(* Logix 5000 project; controller MV vendor 1 type 14 code 217 rev 31.11; software revision 31.00; part 19 of 53 *)
(* tags used below, declared in another part *)
   CheckTimeMask : INT;
   CWD : CHECKWORD_FLAGS;
   Delphi_Does_Eng_Func : BOOL;
   MC_CH1_DR1 : PlantItem;   // CH1_DR1
   MC_CH1_DR2 : PlantItem;   // CH1_DR2
   MC_CH1_DRAIN : PlantItem;   // CH1_DRAIN
   MC_CH1_R1R : PlantItem;   // CH1_R1R
   MC_CH1_R2R : PlantItem;   // CH1_R2R
   MC_CH1_R3R : PlantItem;   // CH1_R3R
   MC_CH1_R4 : PlantItem;   // CH1_R4
   MC_CH1_R4R : PlantItem;   // CH1_R4R
   MC_CH1_R5 : PlantItem;   // CH1_R5
   MC_CH1_R5R : PlantItem;   // CH1_R5R
   MC_CH1_R6 : PlantItem;   // CH1_R6
   MC_CH1_R6R : PlantItem;   // CH1_R6R
   MC_CH1_RR : PlantItem;   // CH1_RR
   MC_N255 : INT[255];   // CHECKWORDS Plant item checkword s
   TempChecktime : DINT;
(* MC_Common, continued *)

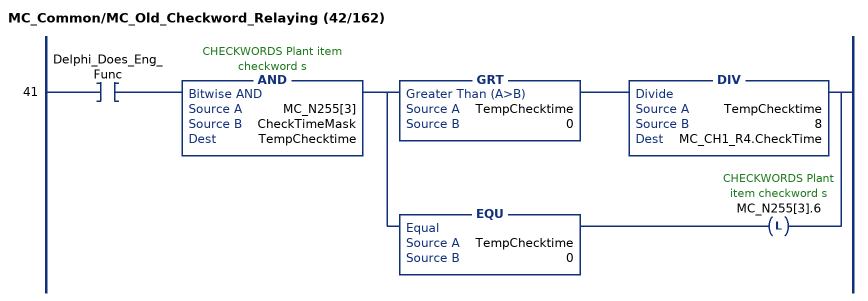
   [picture p312: MC_Common/MC_Old_Checkword_Relaying rungs 41-41]
   41: XIC(Delphi_Does_Eng_Func)AND(MC_N255[3],CheckTimeMask,TempChecktime)[GRT(TempChecktime,0) DIV(TempChecktime,8,MC_CH1_R4.CheckTime) ,EQU(TempChecktime,0) OTL(MC_N255[3].6) ];
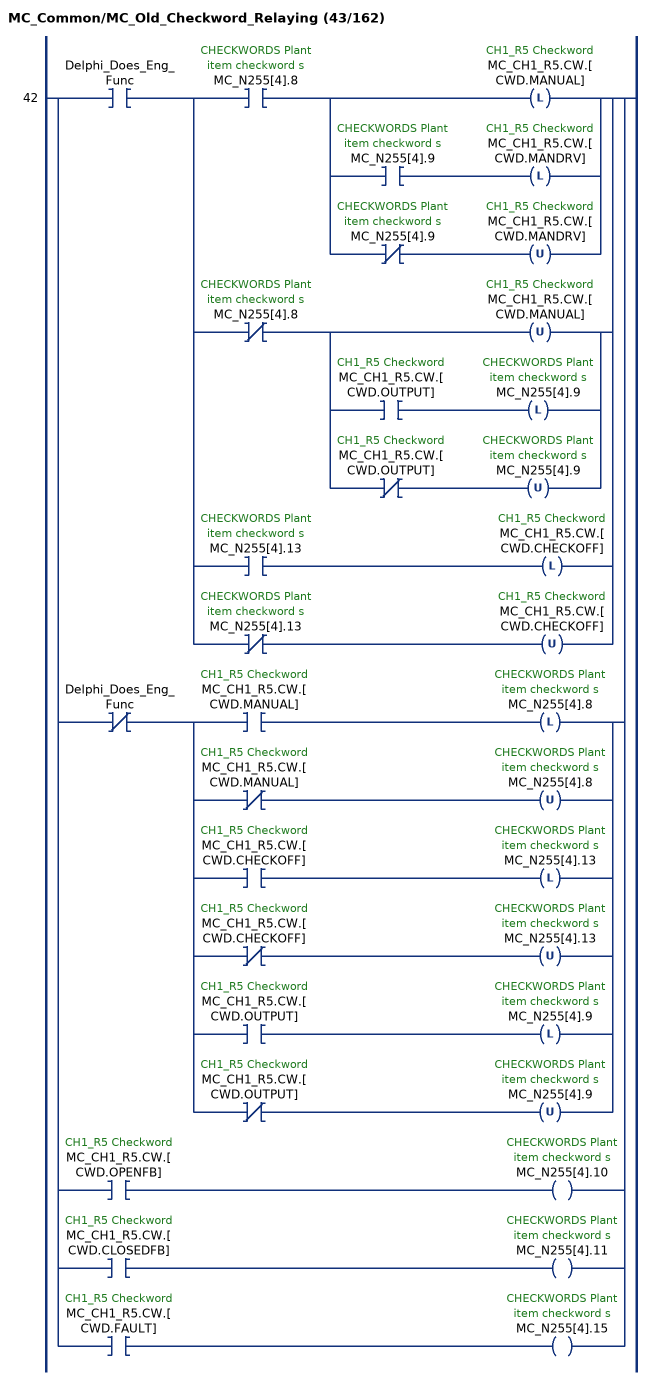
   42: [XIC(Delphi_Does_Eng_Func) [[XIC(MC_N255[4].8) [OTL(MC_CH1_R5.CW.[CWD.MANUAL]) ,XIC(MC_N255[4].9) OTL(MC_CH1_R5.CW.[CWD.MANDRV]) ,XIO(MC_N255[4].9) OTU(MC_CH1_R5.CW.[CWD.MANDRV]) ] ,XIO(MC_N255[4].8) [OTU(MC_CH1_R5.CW.[CWD.MANUAL]) ,[XIC(MC_CH1_R5.CW.[CWD.OUTPUT]) OTL(MC_N255[4].9) ,XIO(MC_CH1_R5.CW.[CWD.OUTPUT]) OTU(MC_N255[4].9) ] ] ] ,[XIC(MC_N255[4].13) OTL(MC_CH1_R5.CW.[CWD.CHECKOFF]) ,XIO(MC_N255[4].13) OTU(MC_CH1_R5.CW.[CWD.CHECKOFF]) ] ] ,XIO(Delphi_Does_Eng_Func) [[XIC(MC_CH1_R5.CW.[CWD.MANUAL]) OTL(MC_N255[4].8) ,XIO(MC_CH1_R5.CW.[CWD.MANUAL]) OTU(MC_N255[4].8) ] ,[XIC(MC_CH1_R5.CW.[CWD.CHECKOFF]) OTL(MC_N255[4].13) ,XIO(MC_CH1_R5.CW.[CWD.CHECKOFF]) OTU(MC_N255[4].13) ] ,[XIC(MC_CH1_R5.CW.[CWD.OUTPUT]) OTL(MC_N255[4].9) ,XIO(MC_CH1_R5.CW.[CWD.OUTPUT]) OTU(MC_N255[4].9) ] ] ,XIC(MC_CH1_R5.CW.[CWD.OPENFB]) OTE(MC_N255[4].10) ,XIC(MC_CH1_R5.CW.[CWD.CLOSEDFB]) OTE(MC_N255[4].11) ,XIC(MC_CH1_R5.CW.[CWD.FAULT]) OTE(MC_N255[4].15) ];
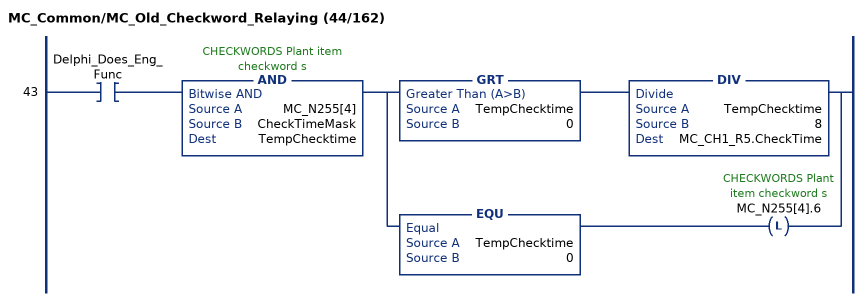
   43: XIC(Delphi_Does_Eng_Func)AND(MC_N255[4],CheckTimeMask,TempChecktime)[GRT(TempChecktime,0) DIV(TempChecktime,8,MC_CH1_R5.CheckTime) ,EQU(TempChecktime,0) OTL(MC_N255[4].6) ];
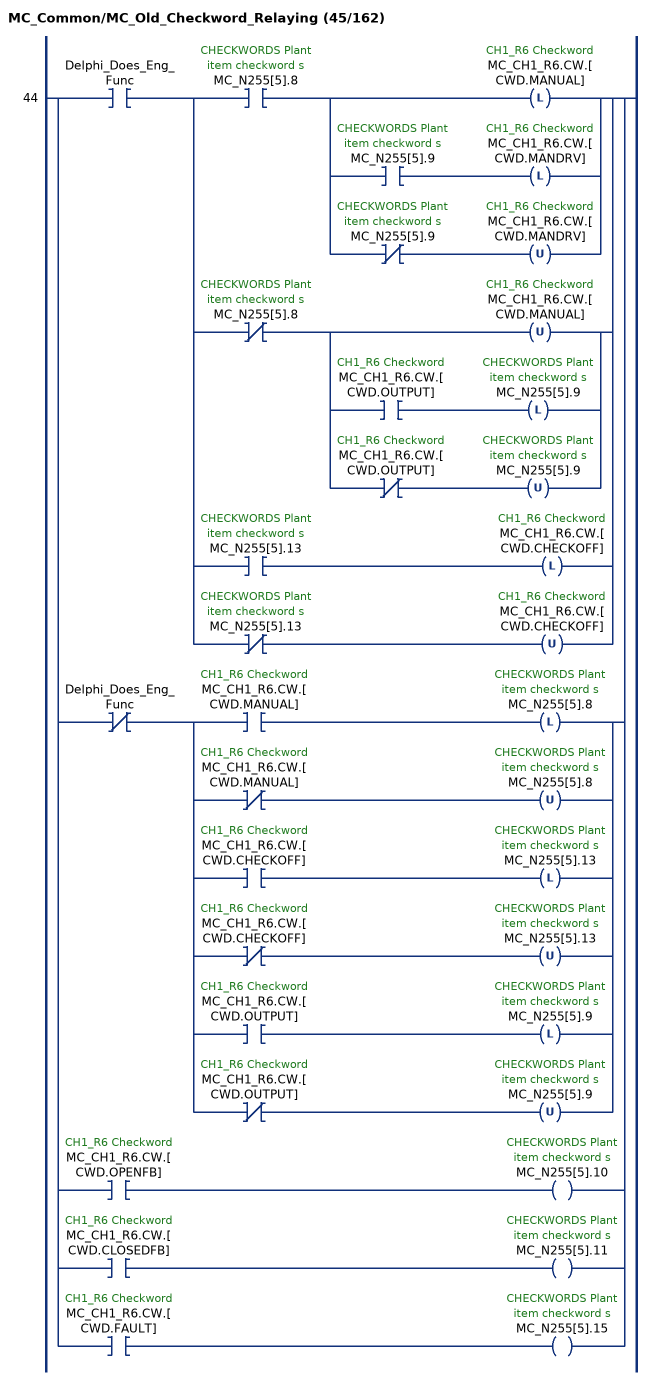
   44: [XIC(Delphi_Does_Eng_Func) [[XIC(MC_N255[5].8) [OTL(MC_CH1_R6.CW.[CWD.MANUAL]) ,XIC(MC_N255[5].9) OTL(MC_CH1_R6.CW.[CWD.MANDRV]) ,XIO(MC_N255[5].9) OTU(MC_CH1_R6.CW.[CWD.MANDRV]) ] ,XIO(MC_N255[5].8) [OTU(MC_CH1_R6.CW.[CWD.MANUAL]) ,[XIC(MC_CH1_R6.CW.[CWD.OUTPUT]) OTL(MC_N255[5].9) ,XIO(MC_CH1_R6.CW.[CWD.OUTPUT]) OTU(MC_N255[5].9) ] ] ] ,[XIC(MC_N255[5].13) OTL(MC_CH1_R6.CW.[CWD.CHECKOFF]) ,XIO(MC_N255[5].13) OTU(MC_CH1_R6.CW.[CWD.CHECKOFF]) ] ] ,XIO(Delphi_Does_Eng_Func) [[XIC(MC_CH1_R6.CW.[CWD.MANUAL]) OTL(MC_N255[5].8) ,XIO(MC_CH1_R6.CW.[CWD.MANUAL]) OTU(MC_N255[5].8) ] ,[XIC(MC_CH1_R6.CW.[CWD.CHECKOFF]) OTL(MC_N255[5].13) ,XIO(MC_CH1_R6.CW.[CWD.CHECKOFF]) OTU(MC_N255[5].13) ] ,[XIC(MC_CH1_R6.CW.[CWD.OUTPUT]) OTL(MC_N255[5].9) ,XIO(MC_CH1_R6.CW.[CWD.OUTPUT]) OTU(MC_N255[5].9) ] ] ,XIC(MC_CH1_R6.CW.[CWD.OPENFB]) OTE(MC_N255[5].10) ,XIC(MC_CH1_R6.CW.[CWD.CLOSEDFB]) OTE(MC_N255[5].11) ,XIC(MC_CH1_R6.CW.[CWD.FAULT]) OTE(MC_N255[5].15) ];
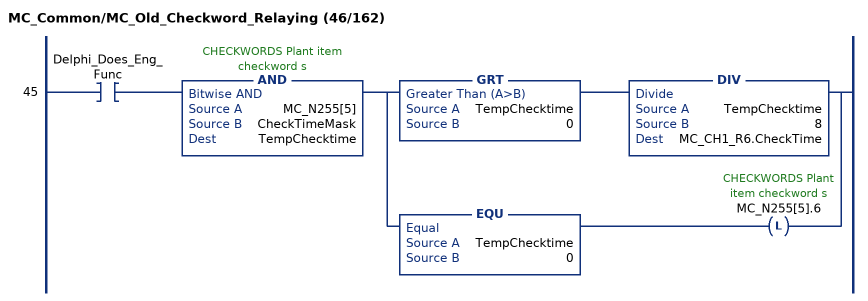
   45: XIC(Delphi_Does_Eng_Func)AND(MC_N255[5],CheckTimeMask,TempChecktime)[GRT(TempChecktime,0) DIV(TempChecktime,8,MC_CH1_R6.CheckTime) ,EQU(TempChecktime,0) OTL(MC_N255[5].6) ];
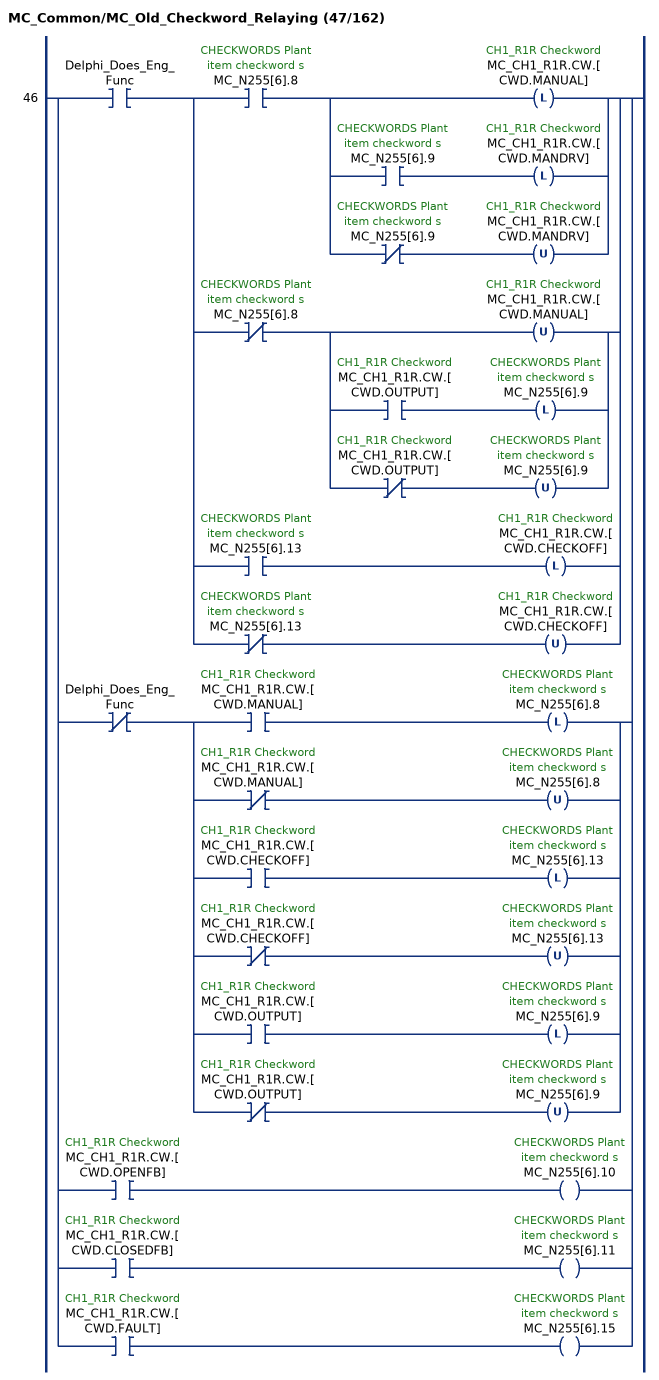
   46: [XIC(Delphi_Does_Eng_Func) [[XIC(MC_N255[6].8) [OTL(MC_CH1_R1R.CW.[CWD.MANUAL]) ,XIC(MC_N255[6].9) OTL(MC_CH1_R1R.CW.[CWD.MANDRV]) ,XIO(MC_N255[6].9) OTU(MC_CH1_R1R.CW.[CWD.MANDRV]) ] ,XIO(MC_N255[6].8) [OTU(MC_CH1_R1R.CW.[CWD.MANUAL]) ,[XIC(MC_CH1_R1R.CW.[CWD.OUTPUT]) OTL(MC_N255[6].9) ,XIO(MC_CH1_R1R.CW.[CWD.OUTPUT]) OTU(MC_N255[6].9) ] ] ] ,[XIC(MC_N255[6].13) OTL(MC_CH1_R1R.CW.[CWD.CHECKOFF]) ,XIO(MC_N255[6].13) OTU(MC_CH1_R1R.CW.[CWD.CHECKOFF]) ] ] ,XIO(Delphi_Does_Eng_Func) [[XIC(MC_CH1_R1R.CW.[CWD.MANUAL]) OTL(MC_N255[6].8) ,XIO(MC_CH1_R1R.CW.[CWD.MANUAL]) OTU(MC_N255[6].8) ] ,[XIC(MC_CH1_R1R.CW.[CWD.CHECKOFF]) OTL(MC_N255[6].13) ,XIO(MC_CH1_R1R.CW.[CWD.CHECKOFF]) OTU(MC_N255[6].13) ] ,[XIC(MC_CH1_R1R.CW.[CWD.OUTPUT]) OTL(MC_N255[6].9) ,XIO(MC_CH1_R1R.CW.[CWD.OUTPUT]) OTU(MC_N255[6].9) ] ] ,XIC(MC_CH1_R1R.CW.[CWD.OPENFB]) OTE(MC_N255[6].10) ,XIC(MC_CH1_R1R.CW.[CWD.CLOSEDFB]) OTE(MC_N255[6].11) ,XIC(MC_CH1_R1R.CW.[CWD.FAULT]) OTE(MC_N255[6].15) ];
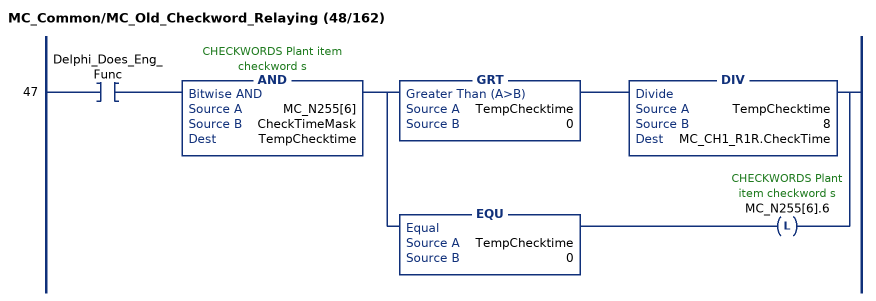
   47: XIC(Delphi_Does_Eng_Func)AND(MC_N255[6],CheckTimeMask,TempChecktime)[GRT(TempChecktime,0) DIV(TempChecktime,8,MC_CH1_R1R.CheckTime) ,EQU(TempChecktime,0) OTL(MC_N255[6].6) ];
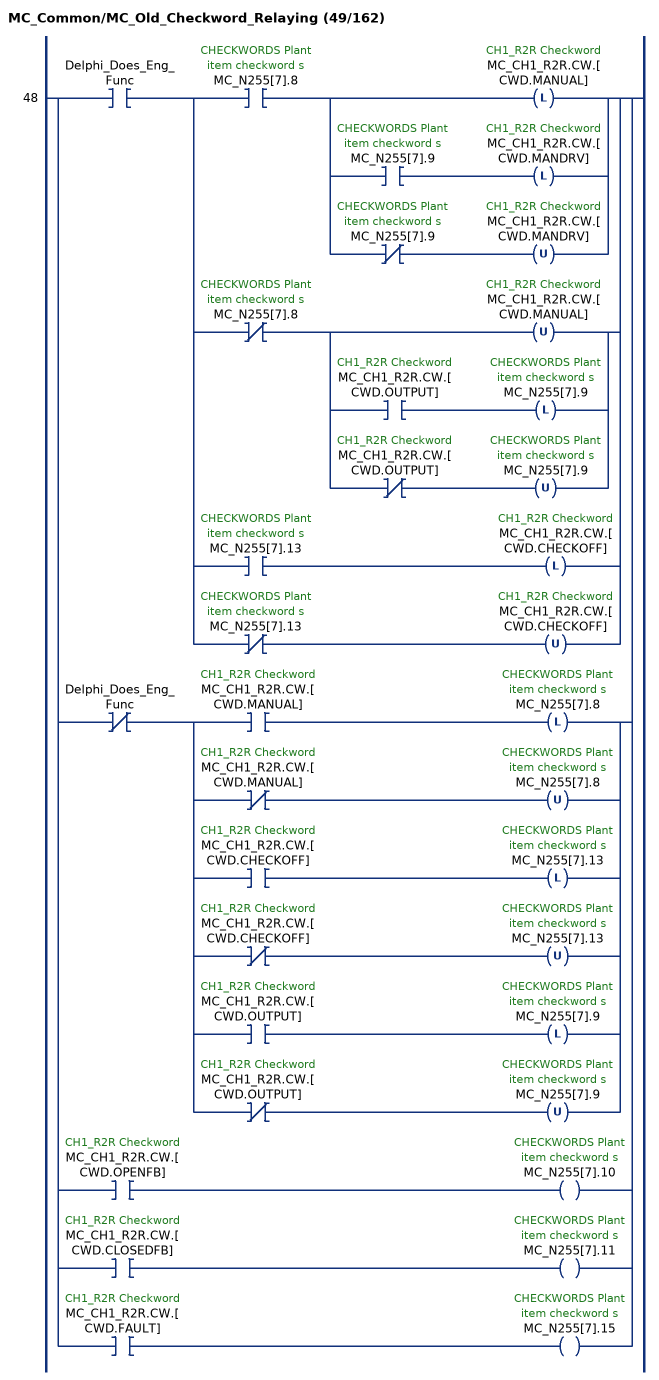
   48: [XIC(Delphi_Does_Eng_Func) [[XIC(MC_N255[7].8) [OTL(MC_CH1_R2R.CW.[CWD.MANUAL]) ,XIC(MC_N255[7].9) OTL(MC_CH1_R2R.CW.[CWD.MANDRV]) ,XIO(MC_N255[7].9) OTU(MC_CH1_R2R.CW.[CWD.MANDRV]) ] ,XIO(MC_N255[7].8) [OTU(MC_CH1_R2R.CW.[CWD.MANUAL]) ,[XIC(MC_CH1_R2R.CW.[CWD.OUTPUT]) OTL(MC_N255[7].9) ,XIO(MC_CH1_R2R.CW.[CWD.OUTPUT]) OTU(MC_N255[7].9) ] ] ] ,[XIC(MC_N255[7].13) OTL(MC_CH1_R2R.CW.[CWD.CHECKOFF]) ,XIO(MC_N255[7].13) OTU(MC_CH1_R2R.CW.[CWD.CHECKOFF]) ] ] ,XIO(Delphi_Does_Eng_Func) [[XIC(MC_CH1_R2R.CW.[CWD.MANUAL]) OTL(MC_N255[7].8) ,XIO(MC_CH1_R2R.CW.[CWD.MANUAL]) OTU(MC_N255[7].8) ] ,[XIC(MC_CH1_R2R.CW.[CWD.CHECKOFF]) OTL(MC_N255[7].13) ,XIO(MC_CH1_R2R.CW.[CWD.CHECKOFF]) OTU(MC_N255[7].13) ] ,[XIC(MC_CH1_R2R.CW.[CWD.OUTPUT]) OTL(MC_N255[7].9) ,XIO(MC_CH1_R2R.CW.[CWD.OUTPUT]) OTU(MC_N255[7].9) ] ] ,XIC(MC_CH1_R2R.CW.[CWD.OPENFB]) OTE(MC_N255[7].10) ,XIC(MC_CH1_R2R.CW.[CWD.CLOSEDFB]) OTE(MC_N255[7].11) ,XIC(MC_CH1_R2R.CW.[CWD.FAULT]) OTE(MC_N255[7].15) ];
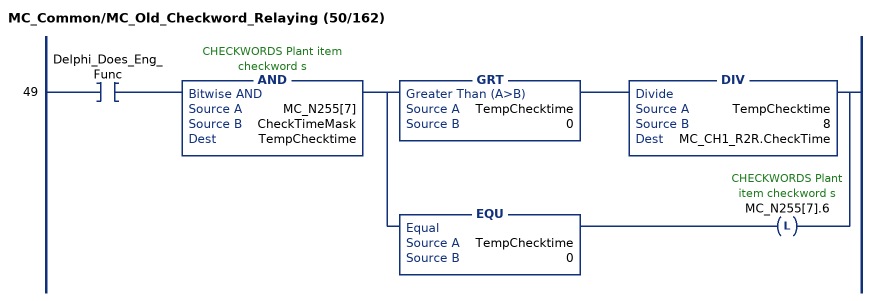
   49: XIC(Delphi_Does_Eng_Func)AND(MC_N255[7],CheckTimeMask,TempChecktime)[GRT(TempChecktime,0) DIV(TempChecktime,8,MC_CH1_R2R.CheckTime) ,EQU(TempChecktime,0) OTL(MC_N255[7].6) ];
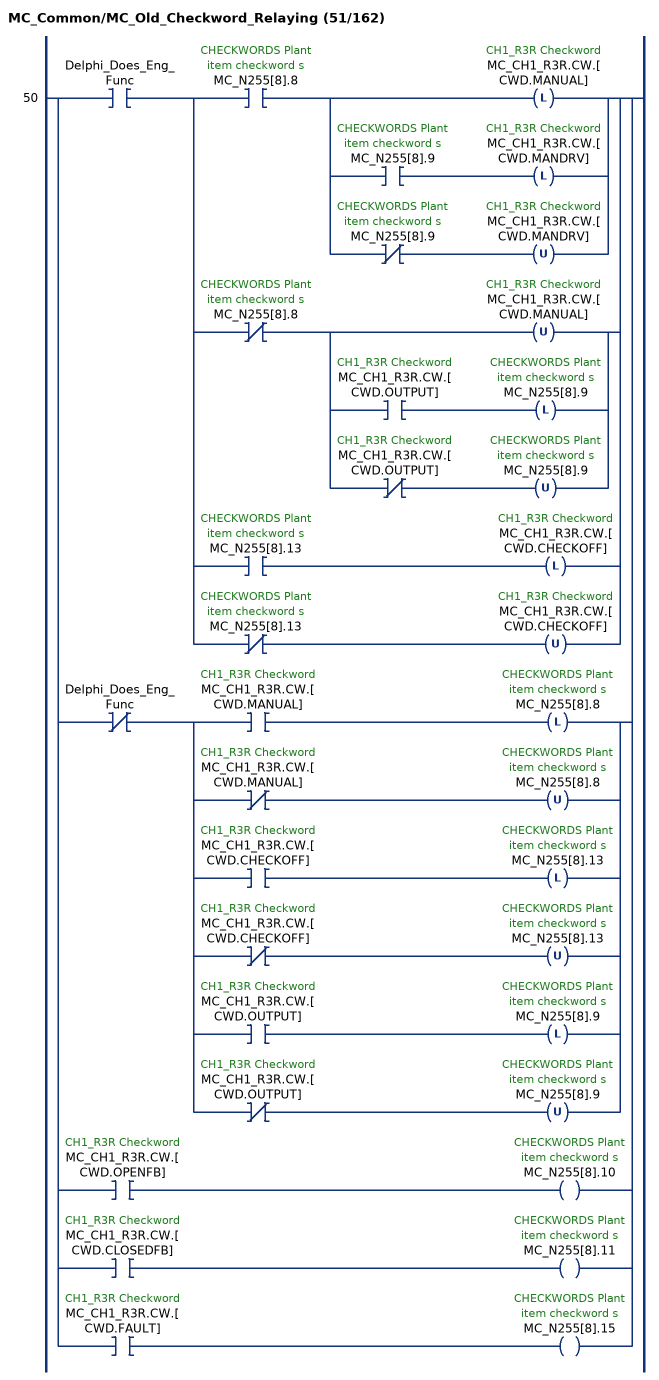
   50: [XIC(Delphi_Does_Eng_Func) [[XIC(MC_N255[8].8) [OTL(MC_CH1_R3R.CW.[CWD.MANUAL]) ,XIC(MC_N255[8].9) OTL(MC_CH1_R3R.CW.[CWD.MANDRV]) ,XIO(MC_N255[8].9) OTU(MC_CH1_R3R.CW.[CWD.MANDRV]) ] ,XIO(MC_N255[8].8) [OTU(MC_CH1_R3R.CW.[CWD.MANUAL]) ,[XIC(MC_CH1_R3R.CW.[CWD.OUTPUT]) OTL(MC_N255[8].9) ,XIO(MC_CH1_R3R.CW.[CWD.OUTPUT]) OTU(MC_N255[8].9) ] ] ] ,[XIC(MC_N255[8].13) OTL(MC_CH1_R3R.CW.[CWD.CHECKOFF]) ,XIO(MC_N255[8].13) OTU(MC_CH1_R3R.CW.[CWD.CHECKOFF]) ] ] ,XIO(Delphi_Does_Eng_Func) [[XIC(MC_CH1_R3R.CW.[CWD.MANUAL]) OTL(MC_N255[8].8) ,XIO(MC_CH1_R3R.CW.[CWD.MANUAL]) OTU(MC_N255[8].8) ] ,[XIC(MC_CH1_R3R.CW.[CWD.CHECKOFF]) OTL(MC_N255[8].13) ,XIO(MC_CH1_R3R.CW.[CWD.CHECKOFF]) OTU(MC_N255[8].13) ] ,[XIC(MC_CH1_R3R.CW.[CWD.OUTPUT]) OTL(MC_N255[8].9) ,XIO(MC_CH1_R3R.CW.[CWD.OUTPUT]) OTU(MC_N255[8].9) ] ] ,XIC(MC_CH1_R3R.CW.[CWD.OPENFB]) OTE(MC_N255[8].10) ,XIC(MC_CH1_R3R.CW.[CWD.CLOSEDFB]) OTE(MC_N255[8].11) ,XIC(MC_CH1_R3R.CW.[CWD.FAULT]) OTE(MC_N255[8].15) ];
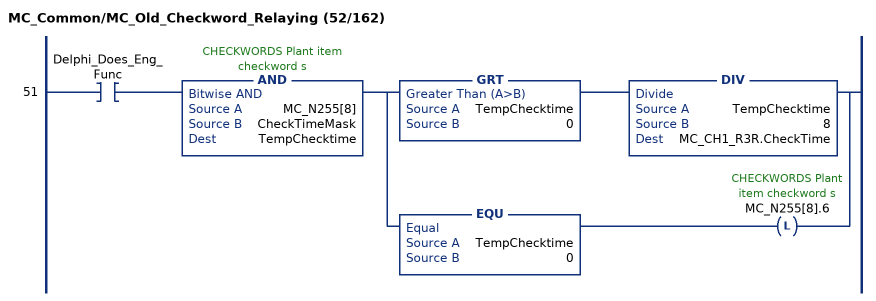
   51: XIC(Delphi_Does_Eng_Func)AND(MC_N255[8],CheckTimeMask,TempChecktime)[GRT(TempChecktime,0) DIV(TempChecktime,8,MC_CH1_R3R.CheckTime) ,EQU(TempChecktime,0) OTL(MC_N255[8].6) ];
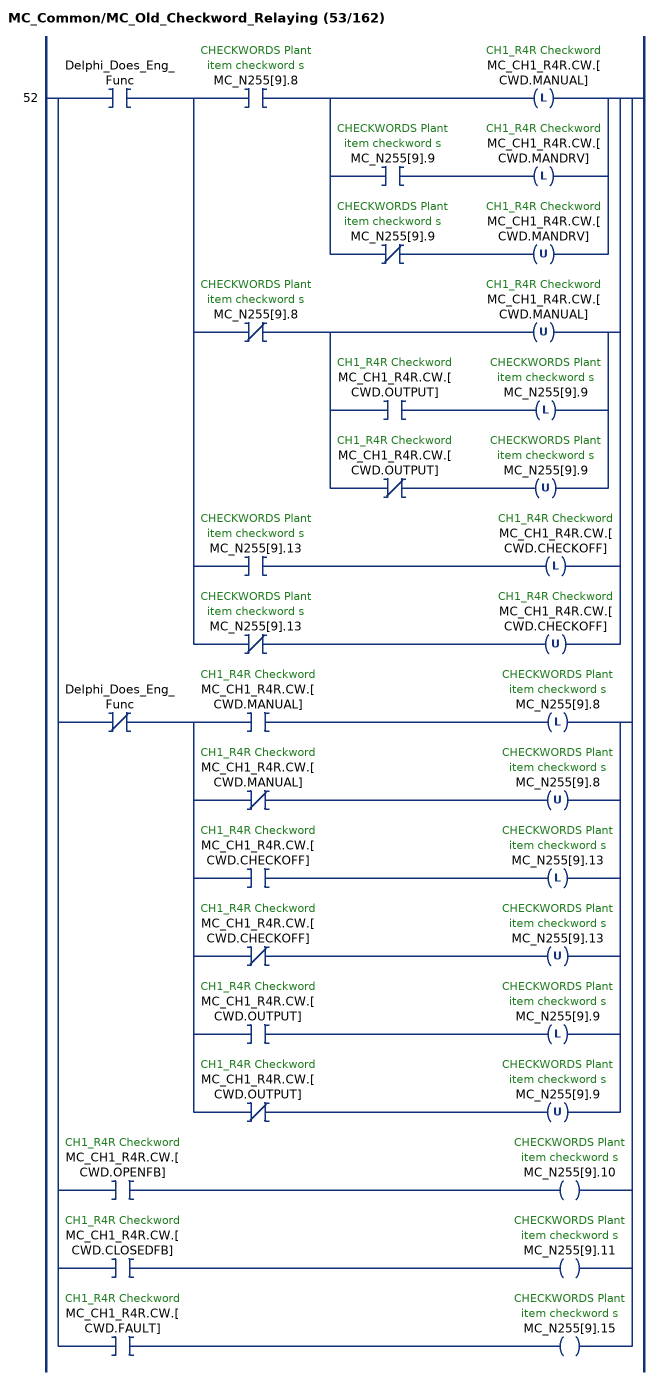
   52: [XIC(Delphi_Does_Eng_Func) [[XIC(MC_N255[9].8) [OTL(MC_CH1_R4R.CW.[CWD.MANUAL]) ,XIC(MC_N255[9].9) OTL(MC_CH1_R4R.CW.[CWD.MANDRV]) ,XIO(MC_N255[9].9) OTU(MC_CH1_R4R.CW.[CWD.MANDRV]) ] ,XIO(MC_N255[9].8) [OTU(MC_CH1_R4R.CW.[CWD.MANUAL]) ,[XIC(MC_CH1_R4R.CW.[CWD.OUTPUT]) OTL(MC_N255[9].9) ,XIO(MC_CH1_R4R.CW.[CWD.OUTPUT]) OTU(MC_N255[9].9) ] ] ] ,[XIC(MC_N255[9].13) OTL(MC_CH1_R4R.CW.[CWD.CHECKOFF]) ,XIO(MC_N255[9].13) OTU(MC_CH1_R4R.CW.[CWD.CHECKOFF]) ] ] ,XIO(Delphi_Does_Eng_Func) [[XIC(MC_CH1_R4R.CW.[CWD.MANUAL]) OTL(MC_N255[9].8) ,XIO(MC_CH1_R4R.CW.[CWD.MANUAL]) OTU(MC_N255[9].8) ] ,[XIC(MC_CH1_R4R.CW.[CWD.CHECKOFF]) OTL(MC_N255[9].13) ,XIO(MC_CH1_R4R.CW.[CWD.CHECKOFF]) OTU(MC_N255[9].13) ] ,[XIC(MC_CH1_R4R.CW.[CWD.OUTPUT]) OTL(MC_N255[9].9) ,XIO(MC_CH1_R4R.CW.[CWD.OUTPUT]) OTU(MC_N255[9].9) ] ] ,XIC(MC_CH1_R4R.CW.[CWD.OPENFB]) OTE(MC_N255[9].10) ,XIC(MC_CH1_R4R.CW.[CWD.CLOSEDFB]) OTE(MC_N255[9].11) ,XIC(MC_CH1_R4R.CW.[CWD.FAULT]) OTE(MC_N255[9].15) ];
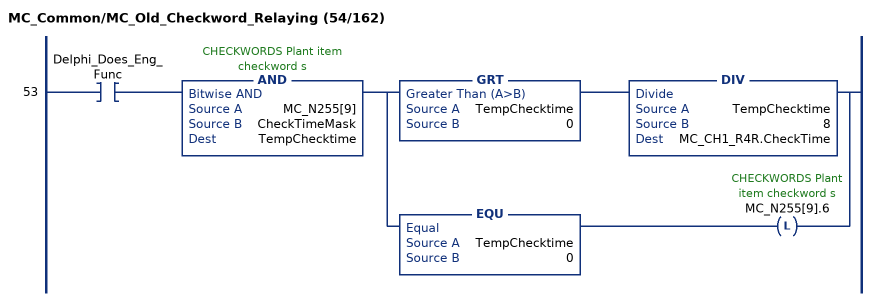
   53: XIC(Delphi_Does_Eng_Func)AND(MC_N255[9],CheckTimeMask,TempChecktime)[GRT(TempChecktime,0) DIV(TempChecktime,8,MC_CH1_R4R.CheckTime) ,EQU(TempChecktime,0) OTL(MC_N255[9].6) ];
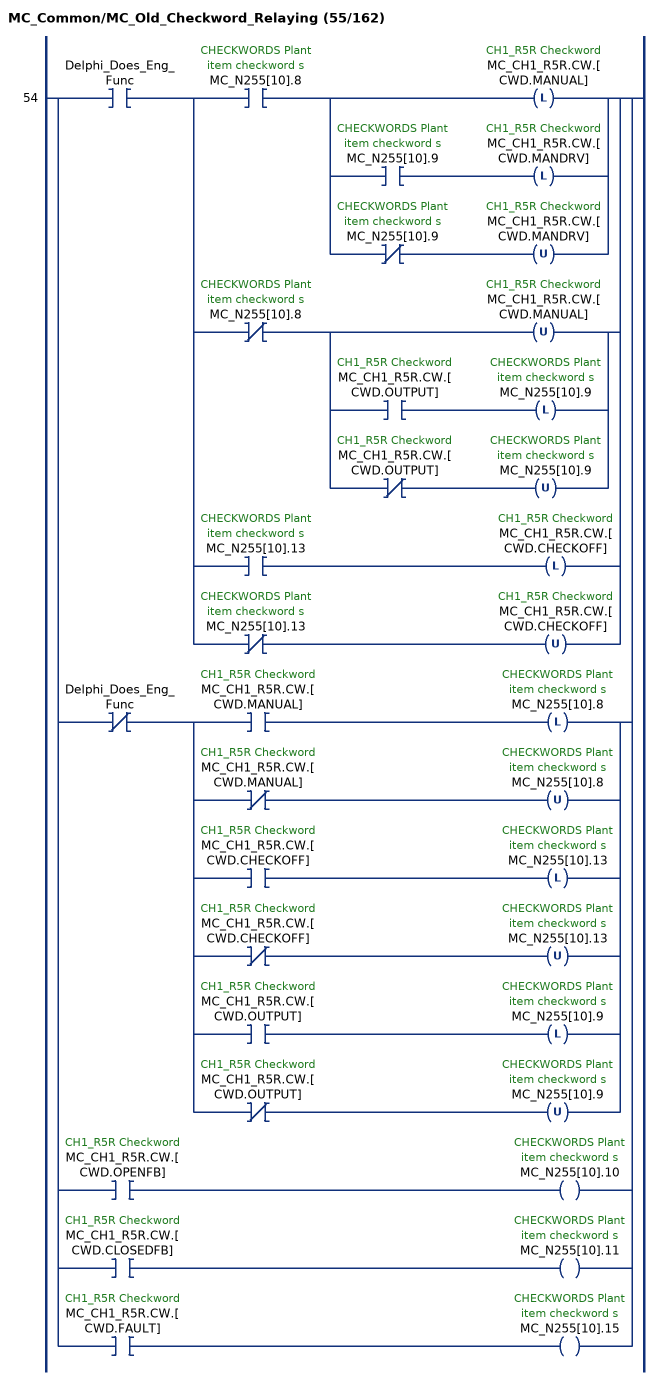
   54: [XIC(Delphi_Does_Eng_Func) [[XIC(MC_N255[10].8) [OTL(MC_CH1_R5R.CW.[CWD.MANUAL]) ,XIC(MC_N255[10].9) OTL(MC_CH1_R5R.CW.[CWD.MANDRV]) ,XIO(MC_N255[10].9) OTU(MC_CH1_R5R.CW.[CWD.MANDRV]) ] ,XIO(MC_N255[10].8) [OTU(MC_CH1_R5R.CW.[CWD.MANUAL]) ,[XIC(MC_CH1_R5R.CW.[CWD.OUTPUT]) OTL(MC_N255[10].9) ,XIO(MC_CH1_R5R.CW.[CWD.OUTPUT]) OTU(MC_N255[10].9) ] ] ] ,[XIC(MC_N255[10].13) OTL(MC_CH1_R5R.CW.[CWD.CHECKOFF]) ,XIO(MC_N255[10].13) OTU(MC_CH1_R5R.CW.[CWD.CHECKOFF]) ] ] ,XIO(Delphi_Does_Eng_Func) [[XIC(MC_CH1_R5R.CW.[CWD.MANUAL]) OTL(MC_N255[10].8) ,XIO(MC_CH1_R5R.CW.[CWD.MANUAL]) OTU(MC_N255[10].8) ] ,[XIC(MC_CH1_R5R.CW.[CWD.CHECKOFF]) OTL(MC_N255[10].13) ,XIO(MC_CH1_R5R.CW.[CWD.CHECKOFF]) OTU(MC_N255[10].13) ] ,[XIC(MC_CH1_R5R.CW.[CWD.OUTPUT]) OTL(MC_N255[10].9) ,XIO(MC_CH1_R5R.CW.[CWD.OUTPUT]) OTU(MC_N255[10].9) ] ] ,XIC(MC_CH1_R5R.CW.[CWD.OPENFB]) OTE(MC_N255[10].10) ,XIC(MC_CH1_R5R.CW.[CWD.CLOSEDFB]) OTE(MC_N255[10].11) ,XIC(MC_CH1_R5R.CW.[CWD.FAULT]) OTE(MC_N255[10].15) ];
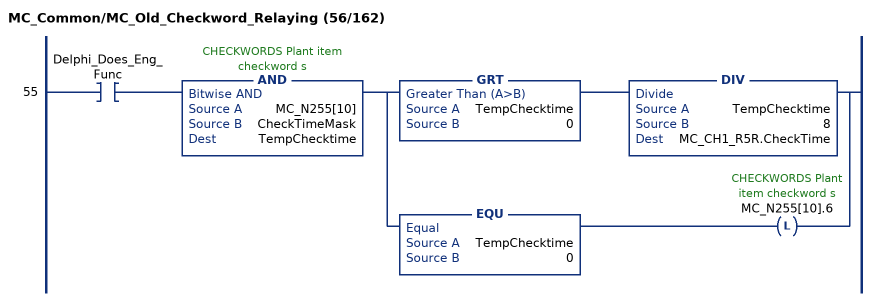
   55: XIC(Delphi_Does_Eng_Func)AND(MC_N255[10],CheckTimeMask,TempChecktime)[GRT(TempChecktime,0) DIV(TempChecktime,8,MC_CH1_R5R.CheckTime) ,EQU(TempChecktime,0) OTL(MC_N255[10].6) ];
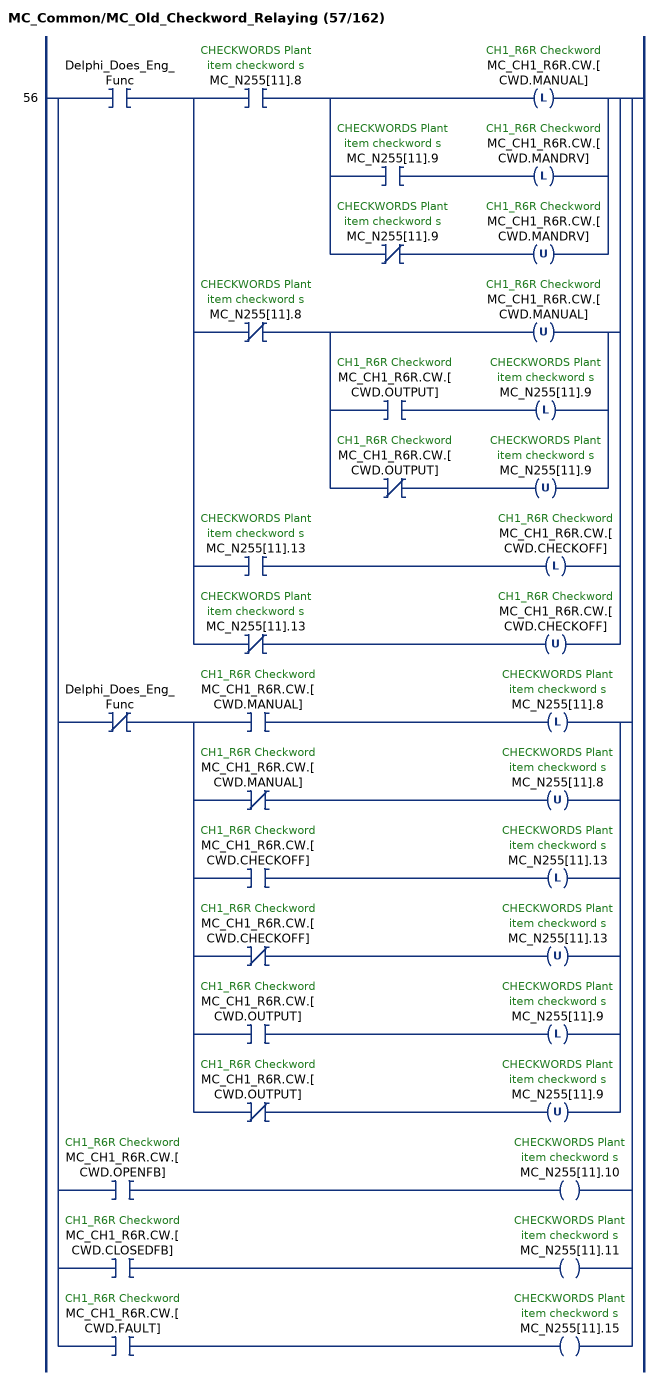
   56: [XIC(Delphi_Does_Eng_Func) [[XIC(MC_N255[11].8) [OTL(MC_CH1_R6R.CW.[CWD.MANUAL]) ,XIC(MC_N255[11].9) OTL(MC_CH1_R6R.CW.[CWD.MANDRV]) ,XIO(MC_N255[11].9) OTU(MC_CH1_R6R.CW.[CWD.MANDRV]) ] ,XIO(MC_N255[11].8) [OTU(MC_CH1_R6R.CW.[CWD.MANUAL]) ,[XIC(MC_CH1_R6R.CW.[CWD.OUTPUT]) OTL(MC_N255[11].9) ,XIO(MC_CH1_R6R.CW.[CWD.OUTPUT]) OTU(MC_N255[11].9) ] ] ] ,[XIC(MC_N255[11].13) OTL(MC_CH1_R6R.CW.[CWD.CHECKOFF]) ,XIO(MC_N255[11].13) OTU(MC_CH1_R6R.CW.[CWD.CHECKOFF]) ] ] ,XIO(Delphi_Does_Eng_Func) [[XIC(MC_CH1_R6R.CW.[CWD.MANUAL]) OTL(MC_N255[11].8) ,XIO(MC_CH1_R6R.CW.[CWD.MANUAL]) OTU(MC_N255[11].8) ] ,[XIC(MC_CH1_R6R.CW.[CWD.CHECKOFF]) OTL(MC_N255[11].13) ,XIO(MC_CH1_R6R.CW.[CWD.CHECKOFF]) OTU(MC_N255[11].13) ] ,[XIC(MC_CH1_R6R.CW.[CWD.OUTPUT]) OTL(MC_N255[11].9) ,XIO(MC_CH1_R6R.CW.[CWD.OUTPUT]) OTU(MC_N255[11].9) ] ] ,XIC(MC_CH1_R6R.CW.[CWD.OPENFB]) OTE(MC_N255[11].10) ,XIC(MC_CH1_R6R.CW.[CWD.CLOSEDFB]) OTE(MC_N255[11].11) ,XIC(MC_CH1_R6R.CW.[CWD.FAULT]) OTE(MC_N255[11].15) ];
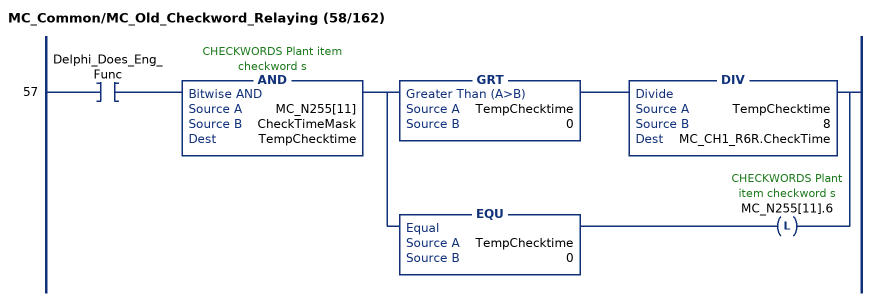
   57: XIC(Delphi_Does_Eng_Func)AND(MC_N255[11],CheckTimeMask,TempChecktime)[GRT(TempChecktime,0) DIV(TempChecktime,8,MC_CH1_R6R.CheckTime) ,EQU(TempChecktime,0) OTL(MC_N255[11].6) ];
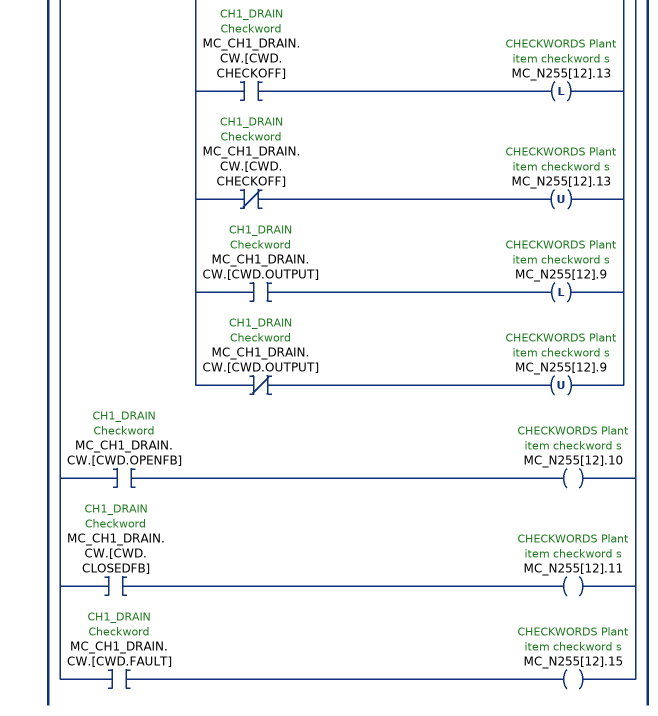
   58: [XIC(Delphi_Does_Eng_Func) [[XIC(MC_N255[12].8) [OTL(MC_CH1_DRAIN.CW.[CWD.MANUAL]) ,XIC(MC_N255[12].9) OTL(MC_CH1_DRAIN.CW.[CWD.MANDRV]) ,XIO(MC_N255[12].9) OTU(MC_CH1_DRAIN.CW.[CWD.MANDRV]) ] ,XIO(MC_N255[12].8) [OTU(MC_CH1_DRAIN.CW.[CWD.MANUAL]) ,[XIC(MC_CH1_DRAIN.CW.[CWD.OUTPUT]) OTL(MC_N255[12].9) ,XIO(MC_CH1_DRAIN.CW.[CWD.OUTPUT]) OTU(MC_N255[12].9) ] ] ] ,[XIC(MC_N255[12].13) OTL(MC_CH1_DRAIN.CW.[CWD.CHECKOFF]) ,XIO(MC_N255[12].13) OTU(MC_CH1_DRAIN.CW.[CWD.CHECKOFF]) ] ] ,XIO(Delphi_Does_Eng_Func) [[XIC(MC_CH1_DRAIN.CW.[CWD.MANUAL]) OTL(MC_N255[12].8) ,XIO(MC_CH1_DRAIN.CW.[CWD.MANUAL]) OTU(MC_N255[12].8) ] ,[XIC(MC_CH1_DRAIN.CW.[CWD.CHECKOFF]) OTL(MC_N255[12].13) ,XIO(MC_CH1_DRAIN.CW.[CWD.CHECKOFF]) OTU(MC_N255[12].13) ] ,[XIC(MC_CH1_DRAIN.CW.[CWD.OUTPUT]) OTL(MC_N255[12].9) ,XIO(MC_CH1_DRAIN.CW.[CWD.OUTPUT]) OTU(MC_N255[12].9) ] ] ,XIC(MC_CH1_DRAIN.CW.[CWD.OPENFB]) OTE(MC_N255[12].10) ,XIC(MC_CH1_DRAIN.CW.[CWD.CLOSEDFB]) OTE(MC_N255[12].11) ,XIC(MC_CH1_DRAIN.CW.[CWD.FAULT]) OTE(MC_N255[12].15) ];
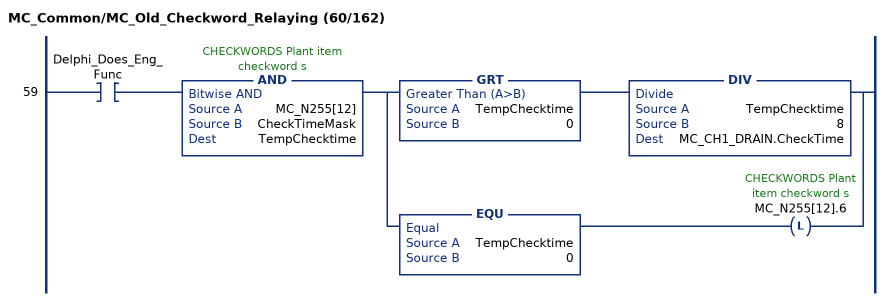
   59: XIC(Delphi_Does_Eng_Func)AND(MC_N255[12],CheckTimeMask,TempChecktime)[GRT(TempChecktime,0) DIV(TempChecktime,8,MC_CH1_DRAIN.CheckTime) ,EQU(TempChecktime,0) OTL(MC_N255[12].6) ];
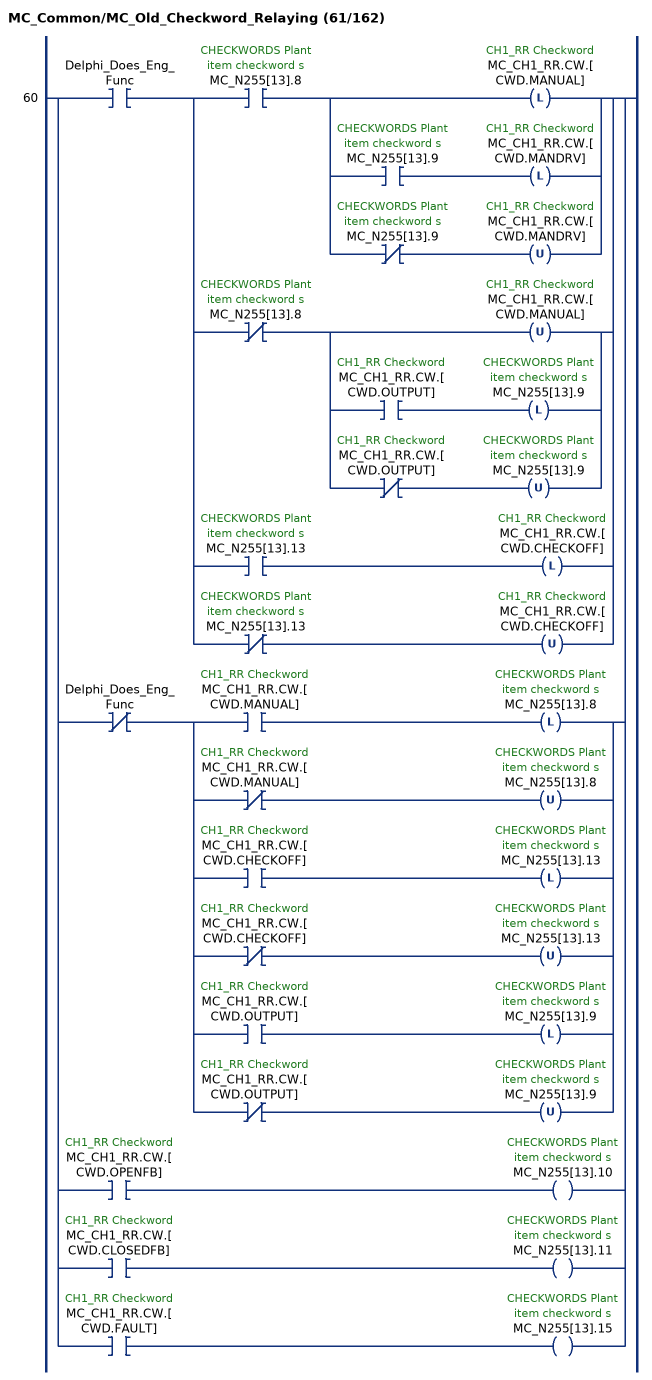
   60: [XIC(Delphi_Does_Eng_Func) [[XIC(MC_N255[13].8) [OTL(MC_CH1_RR.CW.[CWD.MANUAL]) ,XIC(MC_N255[13].9) OTL(MC_CH1_RR.CW.[CWD.MANDRV]) ,XIO(MC_N255[13].9) OTU(MC_CH1_RR.CW.[CWD.MANDRV]) ] ,XIO(MC_N255[13].8) [OTU(MC_CH1_RR.CW.[CWD.MANUAL]) ,[XIC(MC_CH1_RR.CW.[CWD.OUTPUT]) OTL(MC_N255[13].9) ,XIO(MC_CH1_RR.CW.[CWD.OUTPUT]) OTU(MC_N255[13].9) ] ] ] ,[XIC(MC_N255[13].13) OTL(MC_CH1_RR.CW.[CWD.CHECKOFF]) ,XIO(MC_N255[13].13) OTU(MC_CH1_RR.CW.[CWD.CHECKOFF]) ] ] ,XIO(Delphi_Does_Eng_Func) [[XIC(MC_CH1_RR.CW.[CWD.MANUAL]) OTL(MC_N255[13].8) ,XIO(MC_CH1_RR.CW.[CWD.MANUAL]) OTU(MC_N255[13].8) ] ,[XIC(MC_CH1_RR.CW.[CWD.CHECKOFF]) OTL(MC_N255[13].13) ,XIO(MC_CH1_RR.CW.[CWD.CHECKOFF]) OTU(MC_N255[13].13) ] ,[XIC(MC_CH1_RR.CW.[CWD.OUTPUT]) OTL(MC_N255[13].9) ,XIO(MC_CH1_RR.CW.[CWD.OUTPUT]) OTU(MC_N255[13].9) ] ] ,XIC(MC_CH1_RR.CW.[CWD.OPENFB]) OTE(MC_N255[13].10) ,XIC(MC_CH1_RR.CW.[CWD.CLOSEDFB]) OTE(MC_N255[13].11) ,XIC(MC_CH1_RR.CW.[CWD.FAULT]) OTE(MC_N255[13].15) ];
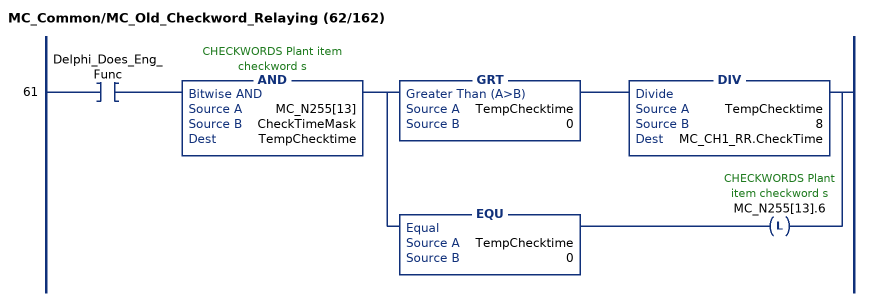
   61: XIC(Delphi_Does_Eng_Func)AND(MC_N255[13],CheckTimeMask,TempChecktime)[GRT(TempChecktime,0) DIV(TempChecktime,8,MC_CH1_RR.CheckTime) ,EQU(TempChecktime,0) OTL(MC_N255[13].6) ];
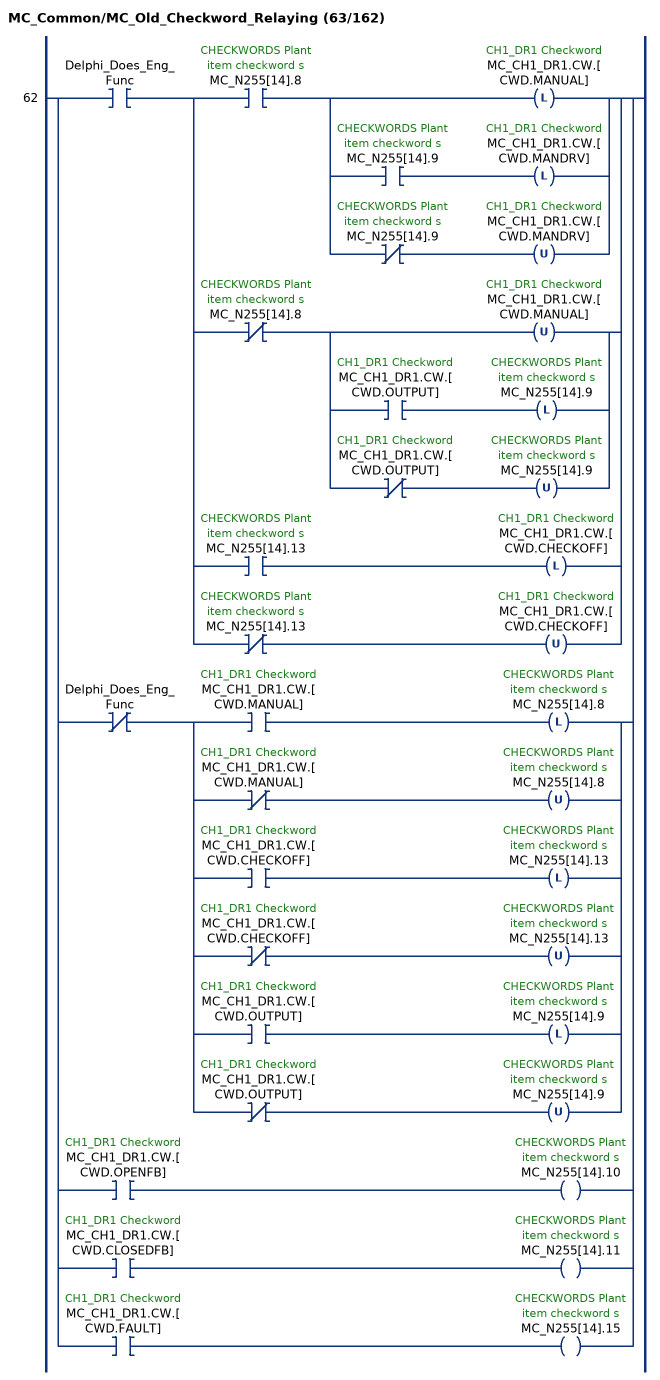
   62: [XIC(Delphi_Does_Eng_Func) [[XIC(MC_N255[14].8) [OTL(MC_CH1_DR1.CW.[CWD.MANUAL]) ,XIC(MC_N255[14].9) OTL(MC_CH1_DR1.CW.[CWD.MANDRV]) ,XIO(MC_N255[14].9) OTU(MC_CH1_DR1.CW.[CWD.MANDRV]) ] ,XIO(MC_N255[14].8) [OTU(MC_CH1_DR1.CW.[CWD.MANUAL]) ,[XIC(MC_CH1_DR1.CW.[CWD.OUTPUT]) OTL(MC_N255[14].9) ,XIO(MC_CH1_DR1.CW.[CWD.OUTPUT]) OTU(MC_N255[14].9) ] ] ] ,[XIC(MC_N255[14].13) OTL(MC_CH1_DR1.CW.[CWD.CHECKOFF]) ,XIO(MC_N255[14].13) OTU(MC_CH1_DR1.CW.[CWD.CHECKOFF]) ] ] ,XIO(Delphi_Does_Eng_Func) [[XIC(MC_CH1_DR1.CW.[CWD.MANUAL]) OTL(MC_N255[14].8) ,XIO(MC_CH1_DR1.CW.[CWD.MANUAL]) OTU(MC_N255[14].8) ] ,[XIC(MC_CH1_DR1.CW.[CWD.CHECKOFF]) OTL(MC_N255[14].13) ,XIO(MC_CH1_DR1.CW.[CWD.CHECKOFF]) OTU(MC_N255[14].13) ] ,[XIC(MC_CH1_DR1.CW.[CWD.OUTPUT]) OTL(MC_N255[14].9) ,XIO(MC_CH1_DR1.CW.[CWD.OUTPUT]) OTU(MC_N255[14].9) ] ] ,XIC(MC_CH1_DR1.CW.[CWD.OPENFB]) OTE(MC_N255[14].10) ,XIC(MC_CH1_DR1.CW.[CWD.CLOSEDFB]) OTE(MC_N255[14].11) ,XIC(MC_CH1_DR1.CW.[CWD.FAULT]) OTE(MC_N255[14].15) ];
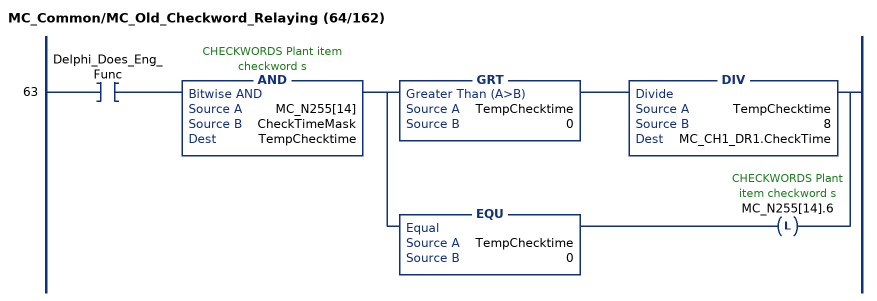
   63: XIC(Delphi_Does_Eng_Func)AND(MC_N255[14],CheckTimeMask,TempChecktime)[GRT(TempChecktime,0) DIV(TempChecktime,8,MC_CH1_DR1.CheckTime) ,EQU(TempChecktime,0) OTL(MC_N255[14].6) ];
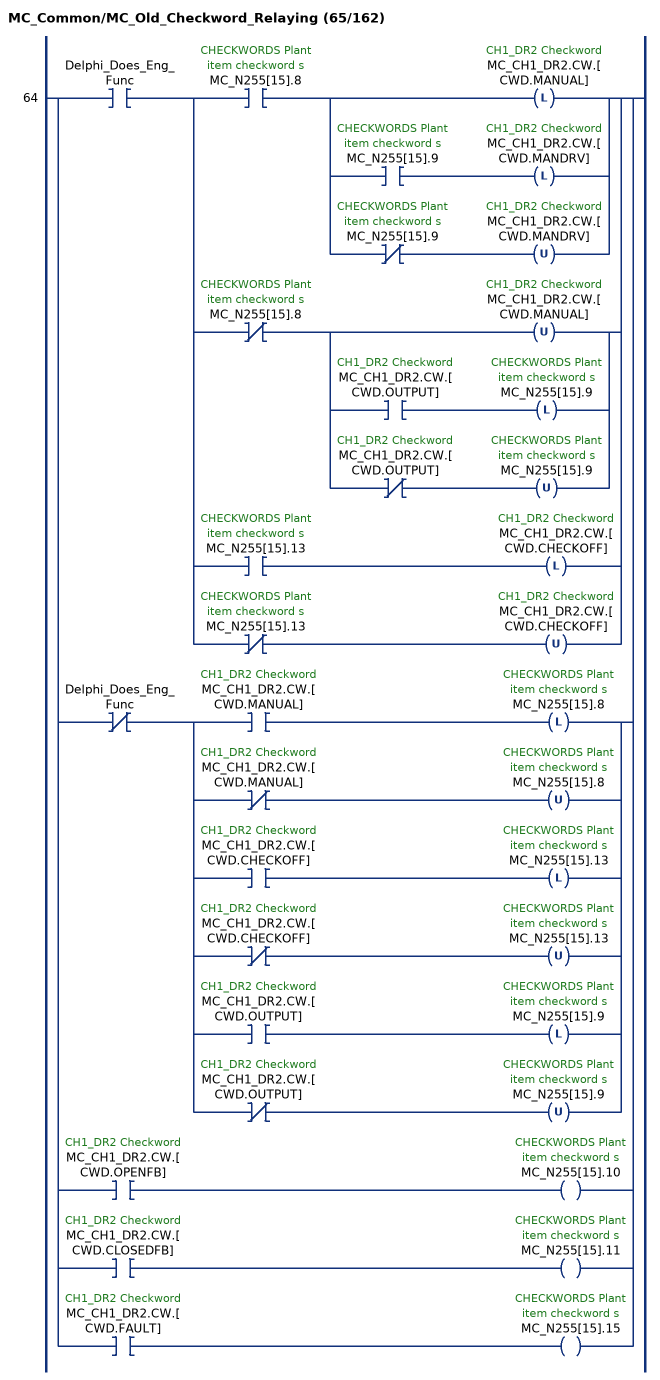
   64: [XIC(Delphi_Does_Eng_Func) [[XIC(MC_N255[15].8) [OTL(MC_CH1_DR2.CW.[CWD.MANUAL]) ,XIC(MC_N255[15].9) OTL(MC_CH1_DR2.CW.[CWD.MANDRV]) ,XIO(MC_N255[15].9) OTU(MC_CH1_DR2.CW.[CWD.MANDRV]) ] ,XIO(MC_N255[15].8) [OTU(MC_CH1_DR2.CW.[CWD.MANUAL]) ,[XIC(MC_CH1_DR2.CW.[CWD.OUTPUT]) OTL(MC_N255[15].9) ,XIO(MC_CH1_DR2.CW.[CWD.OUTPUT]) OTU(MC_N255[15].9) ] ] ] ,[XIC(MC_N255[15].13) OTL(MC_CH1_DR2.CW.[CWD.CHECKOFF]) ,XIO(MC_N255[15].13) OTU(MC_CH1_DR2.CW.[CWD.CHECKOFF]) ] ] ,XIO(Delphi_Does_Eng_Func) [[XIC(MC_CH1_DR2.CW.[CWD.MANUAL]) OTL(MC_N255[15].8) ,XIO(MC_CH1_DR2.CW.[CWD.MANUAL]) OTU(MC_N255[15].8) ] ,[XIC(MC_CH1_DR2.CW.[CWD.CHECKOFF]) OTL(MC_N255[15].13) ,XIO(MC_CH1_DR2.CW.[CWD.CHECKOFF]) OTU(MC_N255[15].13) ] ,[XIC(MC_CH1_DR2.CW.[CWD.OUTPUT]) OTL(MC_N255[15].9) ,XIO(MC_CH1_DR2.CW.[CWD.OUTPUT]) OTU(MC_N255[15].9) ] ] ,XIC(MC_CH1_DR2.CW.[CWD.OPENFB]) OTE(MC_N255[15].10) ,XIC(MC_CH1_DR2.CW.[CWD.CLOSEDFB]) OTE(MC_N255[15].11) ,XIC(MC_CH1_DR2.CW.[CWD.FAULT]) OTE(MC_N255[15].15) ];
